// TIA Portal project "MCP_RB001002" (V15.1) (continued)
   SendWChar[810] := WCHAR#' ';
   SendWChar[811] := WCHAR#' ';
   SendWChar[812] := WCHAR#' ';
   SendWChar[813] := WCHAR#' ';
   SendWChar[814] := WCHAR#' ';
   SendWChar[815] := WCHAR#' ';
   SendWChar[816] := WCHAR#' ';
   SendWChar[817] := WCHAR#' ';
   SendWChar[818] := WCHAR#' ';
   SendWChar[819] := WCHAR#' ';
   SendWChar[820] := WCHAR#' ';
   SendWChar[821] := WCHAR#' ';
   SendWChar[822] := WCHAR#' ';
   SendWChar[823] := WCHAR#' ';
   SendWChar[824] := WCHAR#' ';
   SendWChar[825] := WCHAR#' ';
   SendWChar[826] := WCHAR#' ';
   SendWChar[827] := WCHAR#' ';
   SendWChar[828] := WCHAR#' ';
   SendWChar[829] := WCHAR#' ';
   SendWChar[830] := WCHAR#' ';
   SendWChar[831] := WCHAR#' ';
   SendWChar[832] := WCHAR#' ';
   SendWChar[833] := WCHAR#' ';
   SendWChar[834] := WCHAR#' ';
   SendWChar[835] := WCHAR#' ';
   SendWChar[836] := WCHAR#' ';
   SendWChar[837] := WCHAR#' ';
   SendWChar[838] := WCHAR#' ';
   SendWChar[839] := WCHAR#' ';
   SendWChar[840] := WCHAR#' ';
   SendWChar[841] := WCHAR#' ';
   SendWChar[842] := WCHAR#' ';
   SendWChar[843] := WCHAR#' ';
   SendWChar[844] := WCHAR#' ';
   SendWChar[845] := WCHAR#' ';
   SendWChar[846] := WCHAR#' ';
   SendWChar[847] := WCHAR#' ';
   SendWChar[848] := WCHAR#' ';
   SendWChar[849] := WCHAR#' ';
   SendWChar[850] := WCHAR#' ';
   SendWChar[851] := WCHAR#' ';
   SendWChar[852] := WCHAR#' ';
   SendWChar[853] := WCHAR#' ';
   SendWChar[854] := WCHAR#' ';
   SendWChar[855] := WCHAR#' ';
   SendWChar[856] := WCHAR#' ';
   SendWChar[857] := WCHAR#' ';
   SendWChar[858] := WCHAR#' ';
   SendWChar[859] := WCHAR#' ';
   SendWChar[860] := WCHAR#' ';
   SendWChar[861] := WCHAR#' ';
   SendWChar[862] := WCHAR#' ';
   SendWChar[863] := WCHAR#' ';
   SendWChar[864] := WCHAR#' ';
   SendWChar[865] := WCHAR#' ';
   SendWChar[866] := WCHAR#' ';
   SendWChar[867] := WCHAR#' ';
   SendWChar[868] := WCHAR#' ';
   SendWChar[869] := WCHAR#' ';
   SendWChar[870] := WCHAR#' ';
   SendWChar[871] := WCHAR#' ';
   SendWChar[872] := WCHAR#' ';
   SendWChar[873] := WCHAR#' ';
   SendWChar[874] := WCHAR#' ';
   SendWChar[875] := WCHAR#' ';
   SendWChar[876] := WCHAR#' ';
   SendWChar[877] := WCHAR#' ';
   SendWChar[878] := WCHAR#' ';
   SendWChar[879] := WCHAR#' ';
   SendWChar[880] := WCHAR#' ';
   SendWChar[881] := WCHAR#' ';
   SendWChar[882] := WCHAR#' ';
   SendWChar[883] := WCHAR#' ';
   SendWChar[884] := WCHAR#' ';
   SendWChar[885] := WCHAR#' ';
   SendWChar[886] := WCHAR#' ';
   SendWChar[887] := WCHAR#' ';
   SendWChar[888] := WCHAR#' ';
   SendWChar[889] := WCHAR#' ';
   SendWChar[890] := WCHAR#' ';
   SendWChar[891] := WCHAR#' ';
   SendWChar[892] := WCHAR#' ';
   SendWChar[893] := WCHAR#' ';
   SendWChar[894] := WCHAR#' ';
   SendWChar[895] := WCHAR#' ';
   SendWChar[896] := WCHAR#' ';
   SendWChar[897] := WCHAR#' ';
   SendWChar[898] := WCHAR#' ';
   SendWChar[899] := WCHAR#' ';
   SendWChar[900] := WCHAR#' ';
   SendWChar[901] := WCHAR#' ';
   SendWChar[902] := WCHAR#' ';
   SendWChar[903] := WCHAR#' ';
   SendWChar[904] := WCHAR#' ';
   SendWChar[905] := WCHAR#' ';
   SendWChar[906] := WCHAR#' ';
   SendWChar[907] := WCHAR#' ';
   SendWChar[908] := WCHAR#' ';
   SendWChar[909] := WCHAR#' ';
   SendWChar[910] := WCHAR#' ';
   SendWChar[911] := WCHAR#' ';
   SendWChar[912] := WCHAR#' ';
   SendWChar[913] := WCHAR#' ';
   SendWChar[914] := WCHAR#' ';
   SendWChar[915] := WCHAR#' ';
   SendWChar[916] := WCHAR#' ';
   SendWChar[917] := WCHAR#' ';
   SendWChar[918] := WCHAR#' ';
   SendWChar[919] := WCHAR#' ';
   SendWChar[920] := WCHAR#' ';
   SendWChar[921] := WCHAR#' ';
   SendWChar[922] := WCHAR#' ';
   SendWChar[923] := WCHAR#' ';
   SendWChar[924] := WCHAR#' ';
   SendWChar[925] := WCHAR#' ';
   SendWChar[926] := WCHAR#' ';
   SendWChar[927] := WCHAR#' ';
   SendWChar[928] := WCHAR#' ';
   SendWChar[929] := WCHAR#' ';
   SendWChar[930] := WCHAR#' ';
   SendWChar[931] := WCHAR#' ';
   SendWChar[932] := WCHAR#' ';
   SendWChar[933] := WCHAR#' ';
   SendWChar[934] := WCHAR#' ';
   SendWChar[935] := WCHAR#' ';
   SendWChar[936] := WCHAR#' ';
   SendWChar[937] := WCHAR#' ';
   SendWChar[938] := WCHAR#' ';
   SendWChar[939] := WCHAR#' ';
   SendWChar[940] := WCHAR#' ';
   SendWChar[941] := WCHAR#' ';
   SendWChar[942] := WCHAR#' ';
   SendWChar[943] := WCHAR#' ';
   SendWChar[944] := WCHAR#' ';
   SendWChar[945] := WCHAR#' ';
   SendWChar[946] := WCHAR#' ';
   SendWChar[947] := WCHAR#' ';
   SendWChar[948] := WCHAR#' ';
   SendWChar[949] := WCHAR#' ';
   SendWChar[950] := WCHAR#' ';
   SendWChar[951] := WCHAR#' ';
   SendWChar[952] := WCHAR#' ';
   SendWChar[953] := WCHAR#' ';
   SendWChar[954] := WCHAR#' ';
   SendWChar[955] := WCHAR#' ';
   SendWChar[956] := WCHAR#' ';
   SendWChar[957] := WCHAR#' ';
   SendWChar[958] := WCHAR#' ';
   SendWChar[959] := WCHAR#' ';
   SendWChar[960] := WCHAR#' ';
   SendWChar[961] := WCHAR#' ';
   SendWChar[962] := WCHAR#' ';
   SendWChar[963] := WCHAR#' ';
   SendWChar[964] := WCHAR#' ';
   SendWChar[965] := WCHAR#' ';
   SendWChar[966] := WCHAR#' ';
   SendWChar[967] := WCHAR#' ';
   SendWChar[968] := WCHAR#' ';
   SendWChar[969] := WCHAR#' ';
   SendWChar[970] := WCHAR#' ';
   SendWChar[971] := WCHAR#' ';
   SendWChar[972] := WCHAR#' ';
   SendWChar[973] := WCHAR#' ';
   SendWChar[974] := WCHAR#' ';
   SendWChar[975] := WCHAR#' ';
   SendWChar[976] := WCHAR#' ';
   SendWChar[977] := WCHAR#' ';
   SendWChar[978] := WCHAR#' ';
   SendWChar[979] := WCHAR#' ';
   SendWChar[980] := WCHAR#' ';
   SendWChar[981] := WCHAR#' ';
   SendWChar[982] := WCHAR#' ';
   SendWChar[983] := WCHAR#' ';
   SendWChar[984] := WCHAR#' ';
   SendWChar[985] := WCHAR#' ';
   SendWChar[986] := WCHAR#' ';
   SendWChar[987] := WCHAR#' ';
   SendWChar[988] := WCHAR#' ';
   SendWChar[989] := WCHAR#' ';
   SendWChar[990] := WCHAR#' ';
   SendWChar[991] := WCHAR#' ';
   SendWChar[992] := WCHAR#' ';
   SendWChar[993] := WCHAR#' ';
   SendWChar[994] := WCHAR#' ';
   SendWChar[995] := WCHAR#' ';
   SendWChar[996] := WCHAR#' ';
   SendWChar[997] := WCHAR#' ';
   SendWChar[998] := WCHAR#' ';
   SendWChar[999] := WCHAR#' ';
   SendWChar[1000] := WCHAR#' ';
   SendWChar[1001] := WCHAR#' ';
   SendWChar[1002] := WCHAR#' ';
   SendWChar[1003] := WCHAR#' ';
   SendWChar[1004] := WCHAR#' ';
   SendWChar[1005] := WCHAR#' ';
   SendWChar[1006] := WCHAR#' ';
   SendWChar[1007] := WCHAR#' ';
   SendWChar[1008] := WCHAR#' ';
   SendWChar[1009] := WCHAR#' ';
   SendWChar[1010] := WCHAR#' ';
   SendWChar[1011] := WCHAR#' ';
   SendWChar[1012] := WCHAR#' ';
   SendWChar[1013] := WCHAR#' ';
   SendWChar[1014] := WCHAR#' ';
   SendWChar[1015] := WCHAR#' ';
   SendWChar[1016] := WCHAR#' ';
   SendWChar[1017] := WCHAR#' ';
   SendWChar[1018] := WCHAR#' ';
   SendWChar[1019] := WCHAR#' ';
   SendWChar[1020] := WCHAR#' ';
   SendWChar[1021] := WCHAR#' ';
   SendWChar[1022] := WCHAR#' ';
   SendWChar[1023] := WCHAR#' ';
   SendWChar[1024] := WCHAR#' ';
   SendWChar[1025] := WCHAR#' ';
   SendWChar[1026] := WCHAR#' ';
   SendWChar[1027] := WCHAR#' ';
   SendWChar[1028] := WCHAR#' ';
   SendWChar[1029] := WCHAR#' ';
   SendWChar[1030] := WCHAR#' ';
   SendWChar[1031] := WCHAR#' ';
   SendWChar[1032] := WCHAR#' ';
   SendWChar[1033] := WCHAR#' ';
   SendWChar[1034] := WCHAR#' ';
   SendWChar[1035] := WCHAR#' ';
   SendWChar[1036] := WCHAR#' ';
   SendWChar[1037] := WCHAR#' ';
   SendWChar[1038] := WCHAR#' ';
   SendWChar[1039] := WCHAR#' ';
   SendWChar[1040] := WCHAR#' ';
   SendWChar[1041] := WCHAR#' ';
   SendWChar[1042] := WCHAR#' ';
   SendWChar[1043] := WCHAR#' ';
   SendWChar[1044] := WCHAR#' ';
   SendWChar[1045] := WCHAR#' ';
   SendWChar[1046] := WCHAR#' ';
   SendWChar[1047] := WCHAR#' ';
   SendWChar[1048] := WCHAR#' ';
   SendWChar[1049] := WCHAR#' ';
   SendWChar[1050] := WCHAR#' ';
   SendWChar[1051] := WCHAR#' ';
   SendWChar[1052] := WCHAR#' ';
   SendWChar[1053] := WCHAR#' ';
   SendWChar[1054] := WCHAR#' ';
   SendWChar[1055] := WCHAR#' ';
   SendWChar[1056] := WCHAR#' ';
   SendWChar[1057] := WCHAR#' ';
   SendWChar[1058] := WCHAR#' ';
   SendWChar[1059] := WCHAR#' ';
   SendWChar[1060] := WCHAR#' ';
   SendWChar[1061] := WCHAR#' ';
   SendWChar[1062] := WCHAR#' ';
   SendWChar[1063] := WCHAR#' ';
   SendWChar[1064] := WCHAR#' ';
   SendWChar[1065] := WCHAR#' ';
   SendWChar[1066] := WCHAR#' ';
   SendWChar[1067] := WCHAR#' ';
   SendWChar[1068] := WCHAR#' ';
   SendWChar[1069] := WCHAR#' ';
   SendWChar[1070] := WCHAR#' ';
   SendWChar[1071] := WCHAR#' ';
   SendWChar[1072] := WCHAR#' ';
   SendWChar[1073] := WCHAR#' ';
   SendWChar[1074] := WCHAR#' ';
   SendWChar[1075] := WCHAR#' ';
   SendWChar[1076] := WCHAR#' ';
   SendWChar[1077] := WCHAR#' ';
   SendWChar[1078] := WCHAR#' ';
   SendWChar[1079] := WCHAR#' ';
   SendWChar[1080] := WCHAR#' ';
   SendWChar[1081] := WCHAR#' ';
   SendWChar[1082] := WCHAR#' ';
   SendWChar[1083] := WCHAR#' ';
   SendWChar[1084] := WCHAR#' ';
   SendWChar[1085] := WCHAR#' ';
   SendWChar[1086] := WCHAR#' ';
   SendWChar[1087] := WCHAR#' ';
   SendWChar[1088] := WCHAR#' ';
   SendWChar[1089] := WCHAR#' ';
   SendWChar[1090] := WCHAR#' ';
   SendWChar[1091] := WCHAR#' ';
   SendWChar[1092] := WCHAR#' ';
   SendWChar[1093] := WCHAR#' ';
   SendWChar[1094] := WCHAR#' ';
   SendWChar[1095] := WCHAR#' ';
   SendWChar[1096] := WCHAR#' ';
   SendWChar[1097] := WCHAR#' ';
   SendWChar[1098] := WCHAR#' ';
   SendWChar[1099] := WCHAR#' ';
   SendWChar[1100] := WCHAR#' ';
   SendWChar[1101] := WCHAR#' ';
   SendWChar[1102] := WCHAR#' ';
   SendWChar[1103] := WCHAR#' ';
   SendWChar[1104] := WCHAR#' ';
   SendWChar[1105] := WCHAR#' ';
   SendWChar[1106] := WCHAR#' ';
   SendWChar[1107] := WCHAR#' ';
   SendWChar[1108] := WCHAR#' ';
   SendWChar[1109] := WCHAR#' ';
   SendWChar[1110] := WCHAR#' ';
   SendWChar[1111] := WCHAR#' ';
   SendWChar[1112] := WCHAR#' ';
   SendWChar[1113] := WCHAR#' ';
   SendWChar[1114] := WCHAR#' ';
   SendWChar[1115] := WCHAR#' ';
   SendWChar[1116] := WCHAR#' ';
   SendWChar[1117] := WCHAR#' ';
   SendWChar[1118] := WCHAR#' ';
   SendWChar[1119] := WCHAR#' ';
   SendWChar[1120] := WCHAR#' ';
   SendWChar[1121] := WCHAR#' ';
   SendWChar[1122] := WCHAR#' ';
   SendWChar[1123] := WCHAR#' ';
   SendWChar[1124] := WCHAR#' ';
   SendWChar[1125] := WCHAR#' ';
   SendWChar[1126] := WCHAR#' ';
   SendWChar[1127] := WCHAR#' ';
   SendWChar[1128] := WCHAR#' ';
   SendWChar[1129] := WCHAR#' ';
   SendWChar[1130] := WCHAR#' ';
   SendWChar[1131] := WCHAR#' ';
   SendWChar[1132] := WCHAR#' ';
   SendWChar[1133] := WCHAR#' ';
   SendWChar[1134] := WCHAR#' ';
   SendWChar[1135] := WCHAR#' ';
   SendWChar[1136] := WCHAR#' ';
   SendWChar[1137] := WCHAR#' ';
   SendWChar[1138] := WCHAR#' ';
   SendWChar[1139] := WCHAR#' ';
   SendWChar[1140] := WCHAR#' ';
   SendWChar[1141] := WCHAR#' ';
   SendWChar[1142] := WCHAR#' ';
   SendWChar[1143] := WCHAR#' ';
   SendWChar[1144] := WCHAR#' ';
   SendWChar[1145] := WCHAR#' ';
   SendWChar[1146] := WCHAR#' ';
   SendWChar[1147] := WCHAR#' ';
   SendWChar[1148] := WCHAR#' ';
   SendWChar[1149] := WCHAR#' ';
   SendWChar[1150] := WCHAR#' ';
   SendWChar[1151] := WCHAR#' ';
   SendWChar[1152] := WCHAR#' ';
   SendWChar[1153] := WCHAR#' ';
   SendWChar[1154] := WCHAR#' ';
   SendWChar[1155] := WCHAR#' ';
   SendWChar[1156] := WCHAR#' ';
   SendWChar[1157] := WCHAR#' ';
   SendWChar[1158] := WCHAR#' ';
   SendWChar[1159] := WCHAR#' ';
   SendWChar[1160] := WCHAR#' ';
   SendWChar[1161] := WCHAR#' ';
   SendWChar[1162] := WCHAR#' ';
   SendWChar[1163] := WCHAR#' ';
   SendWChar[1164] := WCHAR#' ';
   SendWChar[1165] := WCHAR#' ';
   SendWChar[1166] := WCHAR#' ';
   SendWChar[1167] := WCHAR#' ';
   SendWChar[1168] := WCHAR#' ';
   SendWChar[1169] := WCHAR#' ';
   SendWChar[1170] := WCHAR#' ';
   SendWChar[1171] := WCHAR#' ';
   SendWChar[1172] := WCHAR#' ';
   SendWChar[1173] := WCHAR#' ';
   SendWChar[1174] := WCHAR#' ';
   SendWChar[1175] := WCHAR#' ';
   SendWChar[1176] := WCHAR#' ';
   SendWChar[1177] := WCHAR#' ';
   SendWChar[1178] := WCHAR#' ';
   SendWChar[1179] := WCHAR#' ';
   SendWChar[1180] := WCHAR#' ';
   SendWChar[1181] := WCHAR#' ';
   SendWChar[1182] := WCHAR#' ';
   SendWChar[1183] := WCHAR#' ';
   SendWChar[1184] := WCHAR#' ';
   SendWChar[1185] := WCHAR#' ';
   SendWChar[1186] := WCHAR#' ';
   SendWChar[1187] := WCHAR#' ';
   SendWChar[1188] := WCHAR#' ';
   SendWChar[1189] := WCHAR#' ';
   SendWChar[1190] := WCHAR#' ';
   SendWChar[1191] := WCHAR#' ';
   SendWChar[1192] := WCHAR#' ';
   SendWChar[1193] := WCHAR#' ';
   SendWChar[1194] := WCHAR#' ';
   SendWChar[1195] := WCHAR#' ';
   SendWChar[1196] := WCHAR#' ';
   SendWChar[1197] := WCHAR#' ';
   SendWChar[1198] := WCHAR#' ';
   SendWChar[1199] := WCHAR#' ';
   SendWChar[1200] := WCHAR#' ';
   SendWChar[1201] := WCHAR#' ';
   SendWChar[1202] := WCHAR#' ';
   SendWChar[1203] := WCHAR#' ';
   SendWChar[1204] := WCHAR#' ';
   SendWChar[1205] := WCHAR#' ';
   SendWChar[1206] := WCHAR#' ';
   SendWChar[1207] := WCHAR#' ';
   SendWChar[1208] := WCHAR#' ';
   SendWChar[1209] := WCHAR#' ';
   SendWChar[1210] := WCHAR#' ';
   SendWChar[1211] := WCHAR#' ';
   SendWChar[1212] := WCHAR#' ';
   SendWChar[1213] := WCHAR#' ';
   SendWChar[1214] := WCHAR#' ';
   SendWChar[1215] := WCHAR#' ';
   SendWChar[1216] := WCHAR#' ';
   SendWChar[1217] := WCHAR#' ';
   SendWChar[1218] := WCHAR#' ';
   SendWChar[1219] := WCHAR#' ';
   SendWChar[1220] := WCHAR#' ';
   SendWChar[1221] := WCHAR#' ';
   SendWChar[1222] := WCHAR#' ';
   SendWChar[1223] := WCHAR#' ';
   SendWChar[1224] := WCHAR#' ';
   SendWChar[1225] := WCHAR#' ';
   SendWChar[1226] := WCHAR#' ';
   SendWChar[1227] := WCHAR#' ';
   SendWChar[1228] := WCHAR#' ';
   SendWChar[1229] := WCHAR#' ';
   SendWChar[1230] := WCHAR#' ';
   SendWChar[1231] := WCHAR#' ';
   SendWChar[1232] := WCHAR#' ';
   SendWChar[1233] := WCHAR#' ';
   SendWChar[1234] := WCHAR#' ';
   SendWChar[1235] := WCHAR#' ';
   SendWChar[1236] := WCHAR#' ';
   SendWChar[1237] := WCHAR#' ';
   SendWChar[1238] := WCHAR#' ';
   SendWChar[1239] := WCHAR#' ';
   SendWChar[1240] := WCHAR#' ';
   SendWChar[1241] := WCHAR#' ';
   SendWChar[1242] := WCHAR#' ';
   SendWChar[1243] := WCHAR#' ';
   SendWChar[1244] := WCHAR#' ';
   SendWChar[1245] := WCHAR#' ';
   SendWChar[1246] := WCHAR#' ';
   SendWChar[1247] := WCHAR#' ';
   SendWChar[1248] := WCHAR#' ';
   SendWChar[1249] := WCHAR#' ';
   SendWChar[1250] := WCHAR#' ';
   SendWChar[1251] := WCHAR#' ';
   SendWChar[1252] := WCHAR#' ';
   SendWChar[1253] := WCHAR#' ';
   SendWChar[1254] := WCHAR#' ';
   SendWChar[1255] := WCHAR#' ';
   SendWChar[1256] := WCHAR#' ';
   SendWChar[1257] := WCHAR#' ';
   SendWChar[1258] := WCHAR#' ';
   SendWChar[1259] := WCHAR#' ';
   SendWChar[1260] := WCHAR#' ';
   SendWChar[1261] := WCHAR#' ';
   SendWChar[1262] := WCHAR#' ';
   SendWChar[1263] := WCHAR#' ';
   SendWChar[1264] := WCHAR#' ';
   SendWChar[1265] := WCHAR#' ';
   SendWChar[1266] := WCHAR#' ';
   SendWChar[1267] := WCHAR#' ';
   SendWChar[1268] := WCHAR#' ';
   SendWChar[1269] := WCHAR#' ';
   SendWChar[1270] := WCHAR#' ';
   SendWChar[1271] := WCHAR#' ';
   SendWChar[1272] := WCHAR#' ';
   SendWChar[1273] := WCHAR#' ';
   SendWChar[1274] := WCHAR#' ';
   SendWChar[1275] := WCHAR#' ';
   SendWChar[1276] := WCHAR#' ';
   SendWChar[1277] := WCHAR#' ';
   SendWChar[1278] := WCHAR#' ';
   SendWChar[1279] := WCHAR#' ';
   SendWChar[1280] := WCHAR#' ';
   SendWChar[1281] := WCHAR#' ';
   SendWChar[1282] := WCHAR#' ';
   SendWChar[1283] := WCHAR#' ';
   SendWChar[1284] := WCHAR#' ';
   SendWChar[1285] := WCHAR#' ';
   SendWChar[1286] := WCHAR#' ';
   SendWChar[1287] := WCHAR#' ';
   SendWChar[1288] := WCHAR#' ';
   SendWChar[1289] := WCHAR#' ';
   SendWChar[1290] := WCHAR#' ';
   SendWChar[1291] := WCHAR#' ';
   SendWChar[1292] := WCHAR#' ';
   SendWChar[1293] := WCHAR#' ';
   SendWChar[1294] := WCHAR#' ';
   SendWChar[1295] := WCHAR#' ';
   SendWChar[1296] := WCHAR#' ';
   SendWChar[1297] := WCHAR#' ';
   SendWChar[1298] := WCHAR#' ';
   SendWChar[1299] := WCHAR#' ';
   SendWChar[1300] := WCHAR#' ';
   SendWChar[1301] := WCHAR#' ';
   SendWChar[1302] := WCHAR#' ';
   SendWChar[1303] := WCHAR#' ';
   SendWChar[1304] := WCHAR#' ';
   SendWChar[1305] := WCHAR#' ';
   SendWChar[1306] := WCHAR#' ';
   SendWChar[1307] := WCHAR#' ';
   SendWChar[1308] := WCHAR#' ';
   SendWChar[1309] := WCHAR#' ';
   SendWChar[1310] := WCHAR#' ';
   SendWChar[1311] := WCHAR#' ';
   SendWChar[1312] := WCHAR#' ';
   SendWChar[1313] := WCHAR#' ';
   SendWChar[1314] := WCHAR#' ';
   SendWChar[1315] := WCHAR#' ';
   SendWChar[1316] := WCHAR#' ';
   SendWChar[1317] := WCHAR#' ';
   SendWChar[1318] := WCHAR#' ';
   SendWChar[1319] := WCHAR#' ';
   SendWChar[1320] := WCHAR#' ';
   SendWChar[1321] := WCHAR#' ';
   SendWChar[1322] := WCHAR#' ';
   SendWChar[1323] := WCHAR#' ';
   SendWChar[1324] := WCHAR#' ';
   SendWChar[1325] := WCHAR#' ';
   SendWChar[1326] := WCHAR#' ';
   SendWChar[1327] := WCHAR#' ';
   SendWChar[1328] := WCHAR#' ';
   SendWChar[1329] := WCHAR#' ';
   SendWChar[1330] := WCHAR#' ';
   SendWChar[1331] := WCHAR#' ';
   SendWChar[1332] := WCHAR#' ';
   SendWChar[1333] := WCHAR#' ';
   SendWChar[1334] := WCHAR#' ';
   SendWChar[1335] := WCHAR#' ';
   SendWChar[1336] := WCHAR#' ';
   SendWChar[1337] := WCHAR#' ';
   SendWChar[1338] := WCHAR#' ';
   SendWChar[1339] := WCHAR#' ';
   SendWChar[1340] := WCHAR#' ';
   SendWChar[1341] := WCHAR#' ';
   SendWChar[1342] := WCHAR#' ';
   SendWChar[1343] := WCHAR#' ';
   SendWChar[1344] := WCHAR#' ';
   SendWChar[1345] := WCHAR#' ';
   SendWChar[1346] := WCHAR#' ';
   SendWChar[1347] := WCHAR#' ';
   SendWChar[1348] := WCHAR#' ';
   SendWChar[1349] := WCHAR#' ';
   SendWChar[1350] := WCHAR#' ';
   SendWChar[1351] := WCHAR#' ';
   SendWChar[1352] := WCHAR#' ';
   SendWChar[1353] := WCHAR#' ';
   SendWChar[1354] := WCHAR#' ';
   SendWChar[1355] := WCHAR#' ';
   SendWChar[1356] := WCHAR#' ';
   SendWChar[1357] := WCHAR#' ';
   SendWChar[1358] := WCHAR#' ';
   SendWChar[1359] := WCHAR#' ';
   SendWChar[1360] := WCHAR#' ';
   SendWChar[1361] := WCHAR#' ';
   SendWChar[1362] := WCHAR#' ';
   SendWChar[1363] := WCHAR#' ';
   SendWChar[1364] := WCHAR#' ';
   SendWChar[1365] := WCHAR#' ';
   SendWChar[1366] := WCHAR#' ';
   SendWChar[1367] := WCHAR#' ';
   SendWChar[1368] := WCHAR#' ';
   SendWChar[1369] := WCHAR#' ';
   SendWChar[1370] := WCHAR#' ';
   SendWChar[1371] := WCHAR#' ';
   SendWChar[1372] := WCHAR#' ';
   SendWChar[1373] := WCHAR#' ';
   SendWChar[1374] := WCHAR#' ';
   SendWChar[1375] := WCHAR#' ';
   SendWChar[1376] := WCHAR#' ';
   SendWChar[1377] := WCHAR#' ';
   SendWChar[1378] := WCHAR#' ';
   SendWChar[1379] := WCHAR#' ';
   SendWChar[1380] := WCHAR#' ';
   SendWChar[1381] := WCHAR#' ';
   SendWChar[1382] := WCHAR#' ';
   SendWChar[1383] := WCHAR#' ';
   SendWChar[1384] := WCHAR#' ';
   SendWChar[1385] := WCHAR#' ';
   SendWChar[1386] := WCHAR#' ';
   SendWChar[1387] := WCHAR#' ';
   SendWChar[1388] := WCHAR#' ';
   SendWChar[1389] := WCHAR#' ';
   SendWChar[1390] := WCHAR#' ';
   SendWChar[1391] := WCHAR#' ';
   SendWChar[1392] := WCHAR#' ';
   SendWChar[1393] := WCHAR#' ';
   SendWChar[1394] := WCHAR#' ';
   SendWChar[1395] := WCHAR#' ';
   SendWChar[1396] := WCHAR#' ';
   SendWChar[1397] := WCHAR#' ';
   SendWChar[1398] := WCHAR#' ';
   SendWChar[1399] := WCHAR#' ';
   SendWChar[1400] := WCHAR#' ';
   SendWChar[1401] := WCHAR#' ';
   SendWChar[1402] := WCHAR#' ';
   SendWChar[1403] := WCHAR#' ';
   SendWChar[1404] := WCHAR#' ';
   SendWChar[1405] := WCHAR#' ';
   SendWChar[1406] := WCHAR#' ';
   SendWChar[1407] := WCHAR#' ';
   SendWChar[1408] := WCHAR#' ';
   SendWChar[1409] := WCHAR#' ';
   SendWChar[1410] := WCHAR#' ';
   SendWChar[1411] := WCHAR#' ';
   SendWChar[1412] := WCHAR#' ';
   SendWChar[1413] := WCHAR#' ';
   SendWChar[1414] := WCHAR#' ';
   SendWChar[1415] := WCHAR#' ';
   SendWChar[1416] := WCHAR#' ';
   SendWChar[1417] := WCHAR#' ';
   SendWChar[1418] := WCHAR#' ';
   SendWChar[1419] := WCHAR#' ';
   SendWChar[1420] := WCHAR#' ';
   SendWChar[1421] := WCHAR#' ';
   SendWChar[1422] := WCHAR#' ';
   SendWChar[1423] := WCHAR#' ';
   SendWChar[1424] := WCHAR#' ';
   SendWChar[1425] := WCHAR#' ';
   SendWChar[1426] := WCHAR#' ';
   SendWChar[1427] := WCHAR#' ';
   SendWChar[1428] := WCHAR#' ';
   SendWChar[1429] := WCHAR#' ';
   SendWChar[1430] := WCHAR#' ';
   SendWChar[1431] := WCHAR#' ';
   SendWChar[1432] := WCHAR#' ';
   SendWChar[1433] := WCHAR#' ';
   SendWChar[1434] := WCHAR#' ';
   SendWChar[1435] := WCHAR#' ';
   SendWChar[1436] := WCHAR#' ';
   SendWChar[1437] := WCHAR#' ';
   SendWChar[1438] := WCHAR#' ';
   SendWChar[1439] := WCHAR#' ';
   SendWChar[1440] := WCHAR#' ';
   SendWChar[1441] := WCHAR#' ';
   SendWChar[1442] := WCHAR#' ';
   SendWChar[1443] := WCHAR#' ';
   SendWChar[1444] := WCHAR#' ';
   SendWChar[1445] := WCHAR#' ';
   SendWChar[1446] := WCHAR#' ';
   SendWChar[1447] := WCHAR#' ';
   SendWChar[1448] := WCHAR#' ';
   SendWChar[1449] := WCHAR#' ';
   SendWChar[1450] := WCHAR#' ';
   SendWChar[1451] := WCHAR#' ';
   SendWChar[1452] := WCHAR#' ';
   SendWChar[1453] := WCHAR#' ';
   SendWChar[1454] := WCHAR#' ';
   SendWChar[1455] := WCHAR#' ';
   SendWChar[1456] := WCHAR#' ';
   SendWChar[1457] := WCHAR#' ';
   SendWChar[1458] := WCHAR#' ';
   SendWChar[1459] := WCHAR#' ';
   SendWChar[1460] := WCHAR#' ';
   SendWChar[1461] := WCHAR#' ';
   SendWChar[1462] := WCHAR#' ';
   SendWChar[1463] := WCHAR#' ';
   SendWChar[1464] := WCHAR#' ';
   SendWChar[1465] := WCHAR#' ';
   SendWChar[1466] := WCHAR#' ';
   SendWChar[1467] := WCHAR#' ';
   SendWChar[1468] := WCHAR#' ';
   SendWChar[1469] := WCHAR#' ';
   SendWChar[1470] := WCHAR#' ';
   SendWChar[1471] := WCHAR#' ';
   SendWChar[1472] := WCHAR#' ';
   SendWChar[1473] := WCHAR#' ';
   SendWChar[1474] := WCHAR#' ';
   SendWChar[1475] := WCHAR#' ';
   SendWChar[1476] := WCHAR#' ';
   SendWChar[1477] := WCHAR#' ';
   SendWChar[1478] := WCHAR#' ';
   SendWChar[1479] := WCHAR#' ';
   SendWChar[1480] := WCHAR#' ';
   SendWChar[1481] := WCHAR#' ';
   SendWChar[1482] := WCHAR#' ';
   SendWChar[1483] := WCHAR#' ';
   SendWChar[1484] := WCHAR#' ';
   SendWChar[1485] := WCHAR#' ';
   SendWChar[1486] := WCHAR#' ';
   SendWChar[1487] := WCHAR#' ';
   SendWChar[1488] := WCHAR#' ';
   SendWChar[1489] := WCHAR#' ';
   SendWChar[1490] := WCHAR#' ';
   SendWChar[1491] := WCHAR#' ';
   SendWChar[1492] := WCHAR#' ';
   SendWChar[1493] := WCHAR#' ';
   SendWChar[1494] := WCHAR#' ';
   SendWChar[1495] := WCHAR#' ';
   SendWChar[1496] := WCHAR#' ';
   SendWChar[1497] := WCHAR#' ';
   SendWChar[1498] := WCHAR#' ';
   SendWChar[1499] := WCHAR#' ';
   SendWChar[1500] := WCHAR#' ';
   SendWChar[1501] := WCHAR#' ';
   SendWChar[1502] := WCHAR#' ';
   SendWChar[1503] := WCHAR#' ';
   SendWChar[1504] := WCHAR#' ';
   SendWChar[1505] := WCHAR#' ';
   SendWChar[1506] := WCHAR#' ';
   SendWChar[1507] := WCHAR#' ';
   SendWChar[1508] := WCHAR#' ';
   SendWChar[1509] := WCHAR#' ';
   SendWChar[1510] := WCHAR#' ';
   SendWChar[1511] := WCHAR#' ';
   SendWChar[1512] := WCHAR#' ';
   SendWChar[1513] := WCHAR#' ';
   SendWChar[1514] := WCHAR#' ';
   SendWChar[1515] := WCHAR#' ';
   SendWChar[1516] := WCHAR#' ';
   SendWChar[1517] := WCHAR#' ';
   SendWChar[1518] := WCHAR#' ';
   SendWChar[1519] := WCHAR#' ';
   SendWChar[1520] := WCHAR#' ';
   SendWChar[1521] := WCHAR#' ';
   SendWChar[1522] := WCHAR#' ';
   SendWChar[1523] := WCHAR#' ';
   SendWChar[1524] := WCHAR#' ';
   SendWChar[1525] := WCHAR#' ';
   SendWChar[1526] := WCHAR#' ';
   SendWChar[1527] := WCHAR#' ';
   SendWChar[1528] := WCHAR#' ';
   SendWChar[1529] := WCHAR#' ';
   SendWChar[1530] := WCHAR#' ';
   SendWChar[1531] := WCHAR#' ';
   SendWChar[1532] := WCHAR#' ';
   SendWChar[1533] := WCHAR#' ';
   SendWChar[1534] := WCHAR#' ';
   SendWChar[1535] := WCHAR#' ';
   SendWChar[1536] := WCHAR#' ';
   SendWChar[1537] := WCHAR#' ';
   SendWChar[1538] := WCHAR#' ';
   SendWChar[1539] := WCHAR#' ';
   SendWChar[1540] := WCHAR#' ';
   SendWChar[1541] := WCHAR#' ';
   SendWChar[1542] := WCHAR#' ';
   SendWChar[1543] := WCHAR#' ';
   SendWChar[1544] := WCHAR#' ';
   SendWChar[1545] := WCHAR#' ';
   SendWChar[1546] := WCHAR#' ';
   SendWChar[1547] := WCHAR#' ';
   SendWChar[1548] := WCHAR#' ';
   SendWChar[1549] := WCHAR#' ';
   SendWChar[1550] := WCHAR#' ';
   SendWChar[1551] := WCHAR#' ';
   SendWChar[1552] := WCHAR#' ';
   SendWChar[1553] := WCHAR#' ';
   SendWChar[1554] := WCHAR#' ';
   SendWChar[1555] := WCHAR#' ';
   SendWChar[1556] := WCHAR#' ';
   SendWChar[1557] := WCHAR#' ';
   SendWChar[1558] := WCHAR#' ';
   SendWChar[1559] := WCHAR#' ';
   SendWChar[1560] := WCHAR#' ';
   SendWChar[1561] := WCHAR#' ';
   SendWChar[1562] := WCHAR#' ';
   SendWChar[1563] := WCHAR#' ';
   SendWChar[1564] := WCHAR#' ';
   SendWChar[1565] := WCHAR#' ';
   SendWChar[1566] := WCHAR#' ';
   SendWChar[1567] := WCHAR#' ';
   SendWChar[1568] := WCHAR#' ';
   SendWChar[1569] := WCHAR#' ';
   SendWChar[1570] := WCHAR#' ';
   SendWChar[1571] := WCHAR#' ';
   SendWChar[1572] := WCHAR#' ';
   SendWChar[1573] := WCHAR#' ';
   SendWChar[1574] := WCHAR#' ';
   SendWChar[1575] := WCHAR#' ';
   SendWChar[1576] := WCHAR#' ';
   SendWChar[1577] := WCHAR#' ';
   SendWChar[1578] := WCHAR#' ';
   SendWChar[1579] := WCHAR#' ';
   SendWChar[1580] := WCHAR#' ';
   SendWChar[1581] := WCHAR#' ';
   SendWChar[1582] := WCHAR#' ';
   SendWChar[1583] := WCHAR#' ';
   SendWChar[1584] := WCHAR#' ';
   SendWChar[1585] := WCHAR#' ';
   SendWChar[1586] := WCHAR#' ';
   SendWChar[1587] := WCHAR#' ';
   SendWChar[1588] := WCHAR#' ';
   SendWChar[1589] := WCHAR#' ';
   SendWChar[1590] := WCHAR#' ';
   SendWChar[1591] := WCHAR#' ';
   SendWChar[1592] := WCHAR#' ';
   SendWChar[1593] := WCHAR#' ';
   SendWChar[1594] := WCHAR#' ';
   SendWChar[1595] := WCHAR#' ';
   SendWChar[1596] := WCHAR#' ';
   SendWChar[1597] := WCHAR#' ';
   SendWChar[1598] := WCHAR#' ';
   SendWChar[1599] := WCHAR#' ';
   SendWChar[1600] := WCHAR#' ';
   SendWChar[1601] := WCHAR#' ';
   SendWChar[1602] := WCHAR#' ';
   SendWChar[1603] := WCHAR#' ';
   SendWChar[1604] := WCHAR#' ';
   SendWChar[1605] := WCHAR#' ';
   SendWChar[1606] := WCHAR#' ';
   SendWChar[1607] := WCHAR#' ';
   SendWChar[1608] := WCHAR#' ';
   SendWChar[1609] := WCHAR#' ';
   SendWChar[1610] := WCHAR#' ';
   SendWChar[1611] := WCHAR#' ';
   SendWChar[1612] := WCHAR#' ';
   SendWChar[1613] := WCHAR#' ';
   SendWChar[1614] := WCHAR#' ';
   SendWChar[1615] := WCHAR#' ';
   SendWChar[1616] := WCHAR#' ';
   SendWChar[1617] := WCHAR#' ';
   SendWChar[1618] := WCHAR#' ';
   SendWChar[1619] := WCHAR#' ';
   SendWChar[1620] := WCHAR#' ';
   SendWChar[1621] := WCHAR#' ';
   SendWChar[1622] := WCHAR#' ';
   SendWChar[1623] := WCHAR#' ';
   SendWChar[1624] := WCHAR#' ';
   SendWChar[1625] := WCHAR#' ';
   SendWChar[1626] := WCHAR#' ';
   SendWChar[1627] := WCHAR#' ';
   SendWChar[1628] := WCHAR#' ';
   SendWChar[1629] := WCHAR#' ';
   SendWChar[1630] := WCHAR#' ';
   SendWChar[1631] := WCHAR#' ';
   SendWChar[1632] := WCHAR#' ';
   SendWChar[1633] := WCHAR#' ';
   SendWChar[1634] := WCHAR#' ';
   SendWChar[1635] := WCHAR#' ';
   SendWChar[1636] := WCHAR#' ';
   SendWChar[1637] := WCHAR#' ';
   SendWChar[1638] := WCHAR#' ';
   SendWChar[1639] := WCHAR#' ';
   SendWChar[1640] := WCHAR#' ';
   SendWChar[1641] := WCHAR#' ';
   SendWChar[1642] := WCHAR#' ';
   SendWChar[1643] := WCHAR#' ';
   SendWChar[1644] := WCHAR#' ';
   SendWChar[1645] := WCHAR#' ';
   SendWChar[1646] := WCHAR#' ';
   SendWChar[1647] := WCHAR#' ';
   SendWChar[1648] := WCHAR#' ';
   SendWChar[1649] := WCHAR#' ';
   SendWChar[1650] := WCHAR#' ';
   SendWChar[1651] := WCHAR#' ';
   SendWChar[1652] := WCHAR#' ';
   SendWChar[1653] := WCHAR#' ';
   SendWChar[1654] := WCHAR#' ';
   SendWChar[1655] := WCHAR#' ';
   SendWChar[1656] := WCHAR#' ';
   SendWChar[1657] := WCHAR#' ';
   SendWChar[1658] := WCHAR#' ';
   SendWChar[1659] := WCHAR#' ';
   SendWChar[1660] := WCHAR#' ';
   SendWChar[1661] := WCHAR#' ';
   SendWChar[1662] := WCHAR#' ';
   SendWChar[1663] := WCHAR#' ';
   SendWChar[1664] := WCHAR#' ';
   SendWChar[1665] := WCHAR#' ';
   SendWChar[1666] := WCHAR#' ';
   SendWChar[1667] := WCHAR#' ';
   SendWChar[1668] := WCHAR#' ';
   SendWChar[1669] := WCHAR#' ';
   SendWChar[1670] := WCHAR#' ';
   SendWChar[1671] := WCHAR#' ';
   SendWChar[1672] := WCHAR#' ';
   SendWChar[1673] := WCHAR#' ';
   SendWChar[1674] := WCHAR#' ';
   SendWChar[1675] := WCHAR#' ';
   SendWChar[1676] := WCHAR#' ';
   SendWChar[1677] := WCHAR#' ';
   SendWChar[1678] := WCHAR#' ';
   SendWChar[1679] := WCHAR#' ';
   SendWChar[1680] := WCHAR#' ';
   SendWChar[1681] := WCHAR#' ';
   SendWChar[1682] := WCHAR#' ';
   SendWChar[1683] := WCHAR#' ';
   SendWChar[1684] := WCHAR#' ';
   SendWChar[1685] := WCHAR#' ';
   SendWChar[1686] := WCHAR#' ';
   SendWChar[1687] := WCHAR#' ';
   SendWChar[1688] := WCHAR#' ';
   SendWChar[1689] := WCHAR#' ';
   SendWChar[1690] := WCHAR#' ';
   SendWChar[1691] := WCHAR#' ';
   SendWChar[1692] := WCHAR#' ';
   SendWChar[1693] := WCHAR#' ';
   SendWChar[1694] := WCHAR#' ';
   SendWChar[1695] := WCHAR#' ';
   SendWChar[1696] := WCHAR#' ';
   SendWChar[1697] := WCHAR#' ';
   SendWChar[1698] := WCHAR#' ';
   SendWChar[1699] := WCHAR#' ';
   SendWChar[1700] := WCHAR#' ';
   SendWChar[1701] := WCHAR#' ';
   SendWChar[1702] := WCHAR#' ';
   SendWChar[1703] := WCHAR#' ';
   SendWChar[1704] := WCHAR#' ';
   SendWChar[1705] := WCHAR#' ';
   SendWChar[1706] := WCHAR#' ';
   SendWChar[1707] := WCHAR#' ';
   SendWChar[1708] := WCHAR#' ';
   SendWChar[1709] := WCHAR#' ';
   SendWChar[1710] := WCHAR#' ';
   SendWChar[1711] := WCHAR#' ';
   SendWChar[1712] := WCHAR#' ';
   SendWChar[1713] := WCHAR#' ';
   SendWChar[1714] := WCHAR#' ';
   SendWChar[1715] := WCHAR#' ';
   SendWChar[1716] := WCHAR#' ';
   SendWChar[1717] := WCHAR#' ';
   SendWChar[1718] := WCHAR#' ';
   SendWChar[1719] := WCHAR#' ';
   SendWChar[1720] := WCHAR#' ';
   SendWChar[1721] := WCHAR#' ';
   SendWChar[1722] := WCHAR#' ';
   SendWChar[1723] := WCHAR#' ';
   SendWChar[1724] := WCHAR#' ';
   SendWChar[1725] := WCHAR#' ';
   SendWChar[1726] := WCHAR#' ';
   SendWChar[1727] := WCHAR#' ';
   SendWChar[1728] := WCHAR#' ';
   SendWChar[1729] := WCHAR#' ';
   SendWChar[1730] := WCHAR#' ';
   SendWChar[1731] := WCHAR#' ';
   SendWChar[1732] := WCHAR#' ';
   SendWChar[1733] := WCHAR#' ';
   SendWChar[1734] := WCHAR#' ';
   SendWChar[1735] := WCHAR#' ';
   SendWChar[1736] := WCHAR#' ';
   SendWChar[1737] := WCHAR#' ';
   SendWChar[1738] := WCHAR#' ';
   SendWChar[1739] := WCHAR#' ';
   SendWChar[1740] := WCHAR#' ';
   SendWChar[1741] := WCHAR#' ';
   SendWChar[1742] := WCHAR#' ';
   SendWChar[1743] := WCHAR#' ';
   SendWChar[1744] := WCHAR#' ';
   SendWChar[1745] := WCHAR#' ';
   SendWChar[1746] := WCHAR#' ';
   SendWChar[1747] := WCHAR#' ';
   SendWChar[1748] := WCHAR#' ';
   SendWChar[1749] := WCHAR#' ';
   SendWChar[1750] := WCHAR#' ';
   SendWChar[1751] := WCHAR#' ';
   SendWChar[1752] := WCHAR#' ';
   SendWChar[1753] := WCHAR#' ';
   SendWChar[1754] := WCHAR#' ';
   SendWChar[1755] := WCHAR#' ';
   SendWChar[1756] := WCHAR#' ';
   SendWChar[1757] := WCHAR#' ';
   SendWChar[1758] := WCHAR#' ';
   SendWChar[1759] := WCHAR#' ';
   SendWChar[1760] := WCHAR#' ';
   SendWChar[1761] := WCHAR#' ';
   SendWChar[1762] := WCHAR#' ';
   SendWChar[1763] := WCHAR#' ';
   SendWChar[1764] := WCHAR#' ';
   SendWChar[1765] := WCHAR#' ';
   SendWChar[1766] := WCHAR#' ';
   SendWChar[1767] := WCHAR#' ';
   SendWChar[1768] := WCHAR#' ';
   SendWChar[1769] := WCHAR#' ';
   SendWChar[1770] := WCHAR#' ';
   SendWChar[1771] := WCHAR#' ';
   SendWChar[1772] := WCHAR#' ';
   SendWChar[1773] := WCHAR#' ';
   SendWChar[1774] := WCHAR#' ';
   SendWChar[1775] := WCHAR#' ';
   SendWChar[1776] := WCHAR#' ';
   SendWChar[1777] := WCHAR#' ';
   SendWChar[1778] := WCHAR#' ';
   SendWChar[1779] := WCHAR#' ';
   SendWChar[1780] := WCHAR#' ';
   SendWChar[1781] := WCHAR#' ';
   SendWChar[1782] := WCHAR#' ';
   SendWChar[1783] := WCHAR#' ';
   SendWChar[1784] := WCHAR#' ';
   SendWChar[1785] := WCHAR#' ';
   SendWChar[1786] := WCHAR#' ';
   SendWChar[1787] := WCHAR#' ';
   SendWChar[1788] := WCHAR#' ';
   SendWChar[1789] := WCHAR#' ';
   SendWChar[1790] := WCHAR#' ';
   SendWChar[1791] := WCHAR#' ';
   SendWChar[1792] := WCHAR#' ';
   SendWChar[1793] := WCHAR#' ';
   SendWChar[1794] := WCHAR#' ';
   SendWChar[1795] := WCHAR#' ';
   SendWChar[1796] := WCHAR#' ';
   SendWChar[1797] := WCHAR#' ';
   SendWChar[1798] := WCHAR#' ';
   SendWChar[1799] := WCHAR#' ';
   SendWChar[1800] := WCHAR#' ';
   SendWChar[1801] := WCHAR#' ';
   SendWChar[1802] := WCHAR#' ';
   SendWChar[1803] := WCHAR#' ';
   SendWChar[1804] := WCHAR#' ';
   SendWChar[1805] := WCHAR#' ';
   SendWChar[1806] := WCHAR#' ';
   SendWChar[1807] := WCHAR#' ';
   SendWChar[1808] := WCHAR#' ';
   SendWChar[1809] := WCHAR#' ';
   SendWChar[1810] := WCHAR#' ';
   SendWChar[1811] := WCHAR#' ';
   SendWChar[1812] := WCHAR#' ';
   SendWChar[1813] := WCHAR#' ';
   SendWChar[1814] := WCHAR#' ';
   SendWChar[1815] := WCHAR#' ';
   SendWChar[1816] := WCHAR#' ';
   SendWChar[1817] := WCHAR#' ';
   SendWChar[1818] := WCHAR#' ';
   SendWChar[1819] := WCHAR#' ';
   SendWChar[1820] := WCHAR#' ';
   SendWChar[1821] := WCHAR#' ';
   SendWChar[1822] := WCHAR#' ';
   SendWChar[1823] := WCHAR#' ';
   SendWChar[1824] := WCHAR#' ';
   SendWChar[1825] := WCHAR#' ';
   SendWChar[1826] := WCHAR#' ';
   SendWChar[1827] := WCHAR#' ';
   SendWChar[1828] := WCHAR#' ';
   SendWChar[1829] := WCHAR#' ';
   SendWChar[1830] := WCHAR#' ';
   SendWChar[1831] := WCHAR#' ';
   SendWChar[1832] := WCHAR#' ';
   SendWChar[1833] := WCHAR#' ';
   SendWChar[1834] := WCHAR#' ';
   SendWChar[1835] := WCHAR#' ';
   SendWChar[1836] := WCHAR#' ';
   SendWChar[1837] := WCHAR#' ';
   SendWChar[1838] := WCHAR#' ';
   SendWChar[1839] := WCHAR#' ';
   SendWChar[1840] := WCHAR#' ';
   SendWChar[1841] := WCHAR#' ';
   SendWChar[1842] := WCHAR#' ';
   SendWChar[1843] := WCHAR#' ';
   SendWChar[1844] := WCHAR#' ';
   SendWChar[1845] := WCHAR#' ';
   SendWChar[1846] := WCHAR#' ';
   SendWChar[1847] := WCHAR#' ';
   SendWChar[1848] := WCHAR#' ';
   SendWChar[1849] := WCHAR#' ';
   SendWChar[1850] := WCHAR#' ';
   SendWChar[1851] := WCHAR#' ';
   SendWChar[1852] := WCHAR#' ';
   SendWChar[1853] := WCHAR#' ';
   SendWChar[1854] := WCHAR#' ';
   SendWChar[1855] := WCHAR#' ';
   SendWChar[1856] := WCHAR#' ';
   SendWChar[1857] := WCHAR#' ';
   SendWChar[1858] := WCHAR#' ';
   SendWChar[1859] := WCHAR#' ';
   SendWChar[1860] := WCHAR#' ';
   SendWChar[1861] := WCHAR#' ';
   SendWChar[1862] := WCHAR#' ';
   SendWChar[1863] := WCHAR#' ';
   SendWChar[1864] := WCHAR#' ';
   SendWChar[1865] := WCHAR#' ';
   SendWChar[1866] := WCHAR#' ';
   SendWChar[1867] := WCHAR#' ';
   SendWChar[1868] := WCHAR#' ';
   SendWChar[1869] := WCHAR#' ';
   SendWChar[1870] := WCHAR#' ';
   SendWChar[1871] := WCHAR#' ';
   SendWChar[1872] := WCHAR#' ';
   SendWChar[1873] := WCHAR#' ';
   SendWChar[1874] := WCHAR#' ';
   SendWChar[1875] := WCHAR#' ';
   SendWChar[1876] := WCHAR#' ';
   SendWChar[1877] := WCHAR#' ';
   SendWChar[1878] := WCHAR#' ';
   SendWChar[1879] := WCHAR#' ';
   SendWChar[1880] := WCHAR#' ';
   SendWChar[1881] := WCHAR#' ';
   SendWChar[1882] := WCHAR#' ';
   SendWChar[1883] := WCHAR#' ';
   SendWChar[1884] := WCHAR#' ';
   SendWChar[1885] := WCHAR#' ';
   SendWChar[1886] := WCHAR#' ';
   SendWChar[1887] := WCHAR#' ';
   SendWChar[1888] := WCHAR#' ';
   SendWChar[1889] := WCHAR#' ';
   SendWChar[1890] := WCHAR#' ';